   //-------------------------------------------------
   //  Signal enable shot finish
   //-------------------------------------------------
         O(;
   //    u    LastBreakFromExternal    // Signal vom ROBOTER !!!
         A     "DB123_MH_IO_Signals".MH[4].IN.MH_Status.shotactive_MH;
         );
         ON    "DB704_MH_Value".Mixinghead[4].ShotBreak;
         O     "DB123_MH_IO_Signals".MH[4].IN.MH_Manual_Mode;
         S     "EnableFinishShot_MH04";

   //-------------------------------------------------
   // Signal to reset shotrelease
   //-------------------------------------------------
         ON    "DB123_MH_IO_Signals".MH[4].IN.MH_Status.shotactive_MH;
         O     "EnableFinishShot_MH04";
         A     "DB123_MH_IO_Signals".MH[4].IN.MH_Status.shotdone_MH;
         S     "ShotFinishedModul_MH04";
   //-------------------------------------------------
   // Shot release
   //-------------------------------------------------
         A     "DB619_State_MPart".Mixinghead[1].Mixingheadvalve."04";
         AN    "ShotFinishedModul_MH04";
         AN    "DB009_Faults".Fault_State_Grp_1_M1;
         AN    "DB009_Faults".Faults_FKT_Grp_1_M1;
         JCN   SO04;
         L     2#0000_0001;
         L     #ControlBitShot;
         OW;
         T     #ControlBitShot;
   //-------------------------------------------------
   // Shot without Timer
   //-------------------------------------------------
   SO04: CLR;
         JCN   SW04;
         L     2#0000_0010;
         L     #ControlBitShot;
         OW;
         T     #ControlBitShot;
   //-------------------------------------------------
   // Shot with Timer
   //-------------------------------------------------
   SW04: A     "DB619_State_MPart".Mixinghead[1].Mixingheadvalve."04";
         AN    "ShotFinishedModul_MH04";
         AN    "DB009_Faults".Fault_State_Grp_1_M1;
         AN    "DB009_Faults".Faults_FKT_Grp_1_M1;
         JCN   SP04;
         L     2#0000_0100;
         L     #ControlBitShot;
         OW;
         T     #ControlBitShot;
   //-----------------------------------------------------------------
   // Service / Production
   //-----------------------------------------------------------------
   SP04: NOP   0;
         A(;
         ON    #TempShotWithMaterial_M1;
         ON    "DB619_State_MPart".MH_at_Machine[1]."04";
         );
         A(;
         ON    #TempShotWithMaterial_M2;
         ON    "DB619_State_MPart".MH_at_Machine[2]."04";
         );
         ON    "DB614_MH_State".MH_Status[4].Switch_Service_ON_OFF;
         JCN   RF03;
         L     2#0000_1000;
         L     #ControlBitShot;
         OW;
         T     #ControlBitShot;
   //-----------------------------------------------------------------
   // Spare Bit 4..6
   //-----------------------------------------------------------------

   //-----------------------------------------------------------------
   // Reset faults
   //-----------------------------------------------------------------
   RF04: A     "DB009_Faults".HF_Faults_Quit;
         JCN   FE04;
         L     2#1000_0000;
         L     #ControlBitShot;
         OW;
         T     #ControlBitShot;

   FE04: NOP   0;
   //-----------------------------------------------------------------
   // Write Output MH Status
   //-----------------------------------------------------------------
         L     "PN_Mixinghead".Mixinghead[4].Digital.Address;
         L     4;
         +D;
         SLD   3;
         LAR1;
         L     #ControlBitShot;
         T     PQB [ AR1 , P#0.0 ];
   //*****************************************************************
   // Cleaning Piston control of mixing head
   //*****************************************************************
         O(;
         L     "PN_Mixinghead".Mixinghead[4].ReinigungskolbenDigital.Address;
         L     0;
         ==I;
         );
         ON    "PN_Mixinghead".Mixinghead[4].ReinigungskolbenDigital.Active;
         JC    em04;

         L     0;
         T     #ControlBitCP;
   //-------------------------------------------------
   // Request cleaning piston after shot
   //-------------------------------------------------
         A     "DB619_State_MPart".ShotMa[1].ShotData.CP_AfterShot;
   //    U     "DB704_MH_Value".Mixinghead[4].WithCleaningPiston
         JCN   CF04;
         L     2#0000_0001;
         L     #ControlBitCP;
         OW;
         T     #ControlBitCP;
   //-------------------------------------------------
   // Request cleaning piston with button
   //-------------------------------------------------
   CF04: A     "DB614_MH_State".MH_CleaningPiston[4].CP_valve_selected;
         JCN   CM04;
         L     2#0000_0010;
         L     #ControlBitCP;
         OW;
         T     #ControlBitCP;
   //-------------------------------------------------
   // Break forward time
   //-------------------------------------------------
   CM04: NOP   0;
   //-----------------------------------------------------------------
   // Reset faults
   //-----------------------------------------------------------------
         A     "DB009_Faults".HF_Faults_Quit;
         JCN   FC04;
         L     2#0000_1000;
         L     #ControlBitCP;
         OW;
         T     #ControlBitCP;
   //-------------------------------------------------
   FC04: NOP   0;
   //-------------------------------------------------
   // Write Output CP Status
   //-------------------------------------------------
         L     "PN_Mixinghead".Mixinghead[4].ReinigungskolbenDigital.Address;
         SLD   3;
         LAR1;
         L     #ControlBitCP;
         T     PQB [ AR1 , P#0.0 ];
   //-------------------------------------------------
         JU    em04;
   //*****************************************************************
   // Setvalue position of cleaning piston MH 3
   //*****************************************************************
   //      L     "DB896_ConfAnaCP_Contr".AnaCleaningPiston[3].RearPosition
   //      UN    "DB610_State_MPart".Cycle_Ma[1].running
   //      SPB   gap1
   //      L     "DB610_State_MPart".ShotMa[1].ShotValues.CP_ThrottleGap
   //      ITD
   //      DTR
   //      L     "DB604_PV_Mixinghead".Mixinghead[3].CleaningPiston.PV_Conf_ActV.Multiplier
   //      *R
   //      RND
   //      L     "DB604_PV_Mixinghead".Mixinghead[3].CleaningPiston.PV_Conf_ActV.OffsetSignal
   //      ITD
   //      +D
   //gap1: T     #ThrottleGap
   //
   //      L     0
   //      L     "DB1232_ProCanIO_MH".AddressMH[3].Ref_PLC_set_value_CP
   //      <D
   //      SPBN  nz01
   //      SLD   3
   //      LAR1
   //      L     #ThrottleGap
   //      T PAW [ AR1 , P#0.0 ]
   //*****************************************************************
   em04: NOP   0;
END_REGION

REGION Network 11: Mixinghead 5
   //--- mixinghead 5 active at a machine ----------------
         O(;
         L     "DB619_State_MPart".ShotMa[1].ShotData.MH_No;
         L     5;
         ==I;
         );
         O(;
         L     "DB619_State_MPart".ShotMa[2].ShotData.MH_No;
         L     5;
         ==I;
         );
         =     #Temp_MH_Shot_MH05;
         JCN   cr05;

         L     "DB704_MH_Value".Mixinghead[5].Corrvalue;
         T     #Temp_CorrValue;

   // Shottime correction
   cr05: NOP   0;

   //----------------------------------------------------------------
   // Read Shottime for next shot
   //----------------------------------------------------------------
         O     "DB619_State_MPart".Cycle[1].PressurizeTimeRuns;
         O     "DB619_State_MPart".Cycle[1].CtrlChangeTimeRuns;
         A     #Temp_MH_Shot_MH05;
         =     "F_CycleRunningMH05";  // Read corr Shottime

         A     #Temp_MH_Shot_MH05;
         A     "DB619_State_MPart".SWU[1].SWU_OK;
         JCN   om05;

         A     "DB619_State_MPart".Operationmode[1].Operation;
         AN    "DB619_State_MPart".ShotMa[1].ShotData.ShotDisabled;
         =     #Temp_OperationMode;

         AN    "DB619_State_MPart".Cycle[1].running;
         R     "StopShotCorrMH05";
         A     "DB110_Interf_Program_M1".Bits.Stop_Cycle;
         A     "DB619_State_MPart".Cycle[1].running;
         S     "StopShotCorrMH05";

         O     "StopShotCorrMH05";
         O     "DB009_Faults".Fault_State_Grp_1_M1;
         ON    "DB619_State_MPart".Operationmode[1].Controllvoltage;
   //      ON    "DB123_MH_IO_Signals".MH[4].IN.MH_Status.shotdone_MH
         =     #Temp_Error;

         CALL  "FC215_SHOT_ADJUST"
         ( IN_Cycle_running   := "F_CycleRunningMH05",  // "DB610_State_MPart".Cycle_Ma[1].running
           IN_Shot_running    := "M_ShotActive",  // "DB610_State_MPart".Cycle_Ma[1].ShotRuns
           IN_OP_Mode_foaming := #Temp_OperationMode,  // "DB610_State_MPart".Operationmode_Ma[1].Operation
           IN_Error_GRP_1     := #Temp_Error,  // "M1001_FaultLevel_1"
           IN_Tool_no         := "DB619_State_MPart".ToolMa[1].ToolNo,
           IN_PS_no           := "ShotNoNextMa1",  // "DB610_State_MPart".ShotDataMa[1].ShotNo
           IN_Set_Shottime_DB := "DB606_PV_Machine".Machine[1].ShotTime.PV_SetV.Value,
           IN_Actual_Shottime := "DB606_PV_Machine".Machine[1].ShotTime.PV_ActV.Value,
           IN_Corrvalue       := #Temp_CorrValue,
           IN_DB_Shotadjust   := "DB315_ShotadjustS",
           IN_ShotRelease     := "DB619_State_MPart".Cycle[1].Shotrelease,
           IN_MhManual        := 0,  //"DB123_MH_IO_Signals".MH[4].IN.MH_Manual_Mode
           IO_Correct_factor  := "DB614_MH_State".ShotAdjustMH[5].CorrFact,
           IO_PAD_Shottime    := "DB614_MH_State".ShotAdjustMH[5].FoamingTime_ProCan,
           IO_Modul_activ     := "DB614_MH_State".ShotAdjustMH[5].ShotCorrActive,
           IO_Helpflag        := "DB614_MH_State".ShotAdjustMH[5].HFShotCorr,
           IO_Last_Shottime   := "DB614_MH_State".ShotAdjustMH[5].LastShottime,
           IO_Soll_for_Corr   := "DB614_MH_State".ShotAdjustMH[5].SetValueForCorr,
           IO_AdrCorrF        := "DB614_MH_State".ShotAdjustMH[5].AdrCorrFact,
           IO_TestProgram     := "DB614_MH_State".ShotAdjustMH[5].ShotCorrTest,
           IO_CorrTimeTest    := "DB614_MH_State".ShotAdjustMH[5].CorrTimeTest
         );

   // Write mixinghead data to procan mudule
   //----------------------------------------------------------------------
   // Check if the communication partner is ready for
   // data transfer to ProCan
   // ---------------------------------------------------------------------
   om05: NOP   0;
         AN    "PN_Mixinghead".Mixinghead[5].Digital.Active;
         AN    "PN_Mixinghead".Mixinghead[5].Analog.Active;
         JC    em05;
   //-----------------------------------------------------------------
   // Output signals of mixing head modul 4
   //-----------------------------------------------------------------
         A     "DB123_MH_IO_Signals".MH[5].OUT.MH.V_SWU_MH;
         =     "V_SWU_MH05";
         A     "DB123_MH_IO_Signals".MH[5].OUT.MH.H_Shotcounter_MH;
         =     "H_Shotcounter_MH05";
         A     "DB123_MH_IO_Signals".MH[5].OUT.MH.V_CP_Forward_MH;
         =     "V_CP_Forward_MH05";
         A     "DB123_MH_IO_Signals".MH[5].OUT.MH.H_CP_Back_MH;
         =     "H_CP_Back_MH05";
         A     "DB123_MH_IO_Signals".MH[5].OUT.MH.H_Rel_Foaming_MH;
         =     "H_Rel_Foaming_MH05";
         A     "DB123_MH_IO_Signals".MH[5].OUT.MH.H_HighPressure_MH;
         =     "H_HighPressure_MH05";
         A     "DB123_MH_IO_Signals".MH[5].OUT.MH.K_Fault_MC;
         =     "K_Fault_MC05";
         A     "DB123_MH_IO_Signals".MH[5].OUT.MH.K_ShotEnd_MC;
         =     "K_ShotEnd_MC05";
         A     "DB123_MH_IO_Signals".MH[5].OUT.MH.V_MH;
         =     "V_MH_open_MH05";
         A     "DB123_MH_IO_Signals".MH[5].OUT.MH.V_LowPressure_Circ_MH;
         =     "V_LowPressure_Circ_MH05";

   //------------------------------------------------------------
   //
   //     Activate mixinghead at ProCan  modul
   //
   //------------------------------------------------------------

   //--------------- Mixinghead 5 --------------------------------
         O     #Temp_MH_Shot_MH05;
         JCN   SV05;
   //-----------------------------------------------------------------
   // Transmit calculated shot time to ProCan
   //-----------------------------------------------------------------
         L     0;
         L     "PN_Mixinghead".Mixinghead[5].Digital.Address;
         <>D;
         JCN   SV05;
         SLD   3;
         LAR1;
         L     "DB614_MH_State".ShotAdjustMH[5].FoamingTime_ProCan;
         T     PQD[AR1, P#0.0];
   SV05: NOP   0;

   //*****************************************************************
   // Shot control of mixing head
   //*****************************************************************
         L     0;
         T     #ControlBitShot;
   //--------------------------------------------------
   // Shotcycle finished reset signals
   //--------------------------------------------------
         AN    "DB619_State_MPart".Mixinghead[1].Mixingheadvalve."05";
         R     "ShotFinishedModul_MH05";
         R     "EnableFinishShot_MH05";

   //-------------------------------------------------
   //  Signal enable shot finish
   //-------------------------------------------------
         O(;
   //    u    LastBreakFromExternal    // Signal vom ROBOTER !!!
         A     "DB123_MH_IO_Signals".MH[5].IN.MH_Status.shotactive_MH;
         );
         ON    "DB704_MH_Value".Mixinghead[5].ShotBreak;
         O     "DB123_MH_IO_Signals".MH[5].IN.MH_Manual_Mode;
         S     "EnableFinishShot_MH05";

   //-------------------------------------------------
   // Signal to reset shotrelease
   //-------------------------------------------------
         ON    "DB123_MH_IO_Signals".MH[5].IN.MH_Status.shotactive_MH;
         O     "EnableFinishShot_MH05";
         A     "DB123_MH_IO_Signals".MH[5].IN.MH_Status.shotdone_MH;
         S     "ShotFinishedModul_MH05";
   //-------------------------------------------------
   // Shot release
   //-------------------------------------------------
         A     "DB619_State_MPart".Mixinghead[1].Mixingheadvalve."05";
         AN    "ShotFinishedModul_MH05";
         AN    "DB009_Faults".Fault_State_Grp_1_M1;
         AN    "DB009_Faults".Faults_FKT_Grp_1_M1;
         JCN   SO05;
         L     2#0000_0001;
         L     #ControlBitShot;
         OW;
         T     #ControlBitShot;
   //-------------------------------------------------
   // Shot without Timer
   //-------------------------------------------------
   SO05: CLR;
         JCN   SW05;
         L     2#0000_0010;
         L     #ControlBitShot;
         OW;
         T     #ControlBitShot;
   //-------------------------------------------------
   // Shot with Timer
   //-------------------------------------------------
   SW05: A     "DB619_State_MPart".Mixinghead[1].Mixingheadvalve."05";
         AN    "ShotFinishedModul_MH05";
         AN    "DB009_Faults".Fault_State_Grp_1_M1;
         AN    "DB009_Faults".Faults_FKT_Grp_1_M1;
         JCN   SP05;
         L     2#0000_0100;
         L     #ControlBitShot;
         OW;
         T     #ControlBitShot;
   //-----------------------------------------------------------------
   // Service / Production
   //-----------------------------------------------------------------
   SP05: NOP   0;
         A(;
         ON    #TempShotWithMaterial_M1;
         ON    "DB619_State_MPart".MH_at_Machine[1]."05";
         );
         A(;
         ON    #TempShotWithMaterial_M2;
         ON    "DB619_State_MPart".MH_at_Machine[2]."05";
         );
         ON    "DB614_MH_State".MH_Status[5].Switch_Service_ON_OFF;
         JCN   RF05;
         L     2#0000_1000;
         L     #ControlBitShot;
         OW;
         T     #ControlBitShot;
   //-----------------------------------------------------------------
   // Spare Bit 4..6
   //-----------------------------------------------------------------

   //-----------------------------------------------------------------
   // Reset faults
   //-----------------------------------------------------------------
   RF05: A     "DB009_Faults".HF_Faults_Quit;
         JCN   FE05;
         L     2#1000_0000;
         L     #ControlBitShot;
         OW;
         T     #ControlBitShot;

   FE05: NOP   0;
   //-----------------------------------------------------------------
   // Write Output MH Status
   //-----------------------------------------------------------------
         L     "PN_Mixinghead".Mixinghead[5].Digital.Address;
         L     4;
         +D;
         SLD   3;
         LAR1;
         L     #ControlBitShot;
         T     PQB [ AR1 , P#0.0 ];
   //*****************************************************************
   // Cleaning Piston control of mixing head
   //*****************************************************************
         O(;
         L     "PN_Mixinghead".Mixinghead[5].ReinigungskolbenDigital.Address;
         L     0;
         ==I;
         );
         ON    "PN_Mixinghead".Mixinghead[5].ReinigungskolbenDigital.Active;
         JC    em05;

         L     0;
         T     #ControlBitCP;
   //-------------------------------------------------
   // Request cleaning piston after shot
   //-------------------------------------------------
         A     "DB619_State_MPart".ShotMa[1].ShotData.CP_AfterShot;
   //    U     "DB704_MH_Value".Mixinghead[5].WithCleaningPiston
         JCN   CF03;
         L     2#0000_0001;
         L     #ControlBitCP;
         OW;
         T     #ControlBitCP;
   //-------------------------------------------------
   // Request cleaning piston with button
   //-------------------------------------------------
   CF05: A     "DB614_MH_State".MH_CleaningPiston[5].CP_valve_selected;
         JCN   CM05;
         L     2#0000_0010;
         L     #ControlBitCP;
         OW;
         T     #ControlBitCP;
   //-------------------------------------------------
   // Break forward time
   //-------------------------------------------------
   CM05: NOP   0;
   //-----------------------------------------------------------------
   // Reset faults
   //-----------------------------------------------------------------
         A     "DB009_Faults".HF_Faults_Quit;
         JCN   FC05;
         L     2#0000_1000;
         L     #ControlBitCP;
         OW;
         T     #ControlBitCP;
   //-------------------------------------------------
   FC05: NOP   0;
   //-------------------------------------------------
   // Write Output CP Status
   //-------------------------------------------------
         L     "PN_Mixinghead".Mixinghead[5].ReinigungskolbenDigital.Address;
         SLD   3;
         LAR1;
         L     #ControlBitCP;
         T     PQB [ AR1 , P#0.0 ];
   //-------------------------------------------------
         JU    em05;
   //*****************************************************************
   // Setvalue position of cleaning piston MH 3
   //*****************************************************************
   //      L     "DB896_ConfAnaCP_Contr".AnaCleaningPiston[3].RearPosition
   //      UN    "DB610_State_MPart".Cycle_Ma[1].running
   //      SPB   gap1
   //      L     "DB610_State_MPart".ShotMa[1].ShotValues.CP_ThrottleGap
   //      ITD
   //      DTR
   //      L     "DB604_PV_Mixinghead".Mixinghead[3].CleaningPiston.PV_Conf_ActV.Multiplier
   //      *R
   //      RND
   //      L     "DB604_PV_Mixinghead".Mixinghead[3].CleaningPiston.PV_Conf_ActV.OffsetSignal
   //      ITD
   //      +D
   //gap1: T     #ThrottleGap
   //
   //      L     0
   //      L     "DB1232_ProCanIO_MH".AddressMH[3].Ref_PLC_set_value_CP
   //      <D
   //      SPBN  nz01
   //      SLD   3
   //      LAR1
   //      L     #ThrottleGap
   //      T PAW [ AR1 , P#0.0 ]
   //*****************************************************************
   em05: NOP   0;
END_REGION

REGION Network 12: Mixinghead 6
   //--- mixinghead 6 active at a machine ----------------
         O(;
         L     "DB619_State_MPart".ShotMa[1].ShotData.MH_No;
         L     6;
         ==I;
         );
         O(;
         L     "DB619_State_MPart".ShotMa[2].ShotData.MH_No;
         L     6;
         ==I;
         );
         =     #Temp_MH_Shot_MH06;
         JCN   cr06;

         L     "DB704_MH_Value".Mixinghead[6].Corrvalue;
         T     #Temp_CorrValue;

   // Shottime correction
   cr06: NOP   0;

   //----------------------------------------------------------------
   // Read Shottime for next shot
   //----------------------------------------------------------------
         O     "DB619_State_MPart".Cycle[1].PressurizeTimeRuns;
         O     "DB619_State_MPart".Cycle[1].CtrlChangeTimeRuns;
         A     #Temp_MH_Shot_MH06;
         =     "F_CycleRunningMH06";  // Read corr Shottime

         A     #Temp_MH_Shot_MH06;
         A     "DB619_State_MPart".SWU[1].SWU_OK;
         JCN   om06;

         A     "DB619_State_MPart".Operationmode[1].Operation;
         AN    "DB619_State_MPart".ShotMa[1].ShotData.ShotDisabled;
         =     #Temp_OperationMode;

         AN    "DB619_State_MPart".Cycle[1].running;
         R     "StopShotCorrMH06";
         A     "DB110_Interf_Program_M1".Bits.Stop_Cycle;
         A     "DB619_State_MPart".Cycle[1].running;
         S     "StopShotCorrMH06";

         O     "StopShotCorrMH06";
         O     "DB009_Faults".Fault_State_Grp_1_M1;
         ON    "DB619_State_MPart".Operationmode[1].Controllvoltage;
   //      ON    "DB123_MH_IO_Signals".MH[4].IN.MH_Status.shotdone_MH
         =     #Temp_Error;

         CALL  "FC215_SHOT_ADJUST"
         ( IN_Cycle_running   := "F_CycleRunningMH06",  // "DB610_State_MPart".Cycle_Ma[1].running
           IN_Shot_running    := "M_ShotActive",  // "DB610_State_MPart".Cycle_Ma[1].ShotRuns
           IN_OP_Mode_foaming := #Temp_OperationMode,  // "DB610_State_MPart".Operationmode_Ma[1].Operation
           IN_Error_GRP_1     := #Temp_Error,  // "M1001_FaultLevel_1"
           IN_Tool_no         := "DB619_State_MPart".ToolMa[1].ToolNo,
           IN_PS_no           := "ShotNoNextMa1",  // "DB610_State_MPart".ShotDataMa[1].ShotNo
           IN_Set_Shottime_DB := "DB606_PV_Machine".Machine[1].ShotTime.PV_SetV.Value,
           IN_Actual_Shottime := "DB606_PV_Machine".Machine[1].ShotTime.PV_ActV.Value,
           IN_Corrvalue       := #Temp_CorrValue,
           IN_DB_Shotadjust   := "DB315_ShotadjustS",
           IN_ShotRelease     := "DB619_State_MPart".Cycle[1].Shotrelease,
           IN_MhManual        := 0,  //"DB123_MH_IO_Signals".MH[4].IN.MH_Manual_Mode
           IO_Correct_factor  := "DB614_MH_State".ShotAdjustMH[6].CorrFact,
           IO_PAD_Shottime    := "DB614_MH_State".ShotAdjustMH[6].FoamingTime_ProCan,
           IO_Modul_activ     := "DB614_MH_State".ShotAdjustMH[6].ShotCorrActive,
           IO_Helpflag        := "DB614_MH_State".ShotAdjustMH[6].HFShotCorr,
           IO_Last_Shottime   := "DB614_MH_State".ShotAdjustMH[6].LastShottime,
           IO_Soll_for_Corr   := "DB614_MH_State".ShotAdjustMH[6].SetValueForCorr,
           IO_AdrCorrF        := "DB614_MH_State".ShotAdjustMH[6].AdrCorrFact,
           IO_TestProgram     := "DB614_MH_State".ShotAdjustMH[6].ShotCorrTest,
           IO_CorrTimeTest    := "DB614_MH_State".ShotAdjustMH[6].CorrTimeTest
         );

   // Write mixinghead data to procan mudule
   //----------------------------------------------------------------------
   // Check if the communication partner is ready for
   // data transfer to ProCan
   // ---------------------------------------------------------------------
   om06: NOP   0;
         AN    "PN_Mixinghead".Mixinghead[6].Digital.Active;
         AN    "PN_Mixinghead".Mixinghead[6].Analog.Active;
         JC    em06;
   //-----------------------------------------------------------------
   // Output signals of mixing head modul 6
   //-----------------------------------------------------------------
         A     "DB123_MH_IO_Signals".MH[6].OUT.MH.V_SWU_MH;
         =     "V_SWU_MH06";
         A     "DB123_MH_IO_Signals".MH[6].OUT.MH.H_Shotcounter_MH;
         =     "H_Shotcounter_MH06";
         A     "DB123_MH_IO_Signals".MH[6].OUT.MH.V_CP_Forward_MH;
         =     "V_CP_Forward_MH06";
         A     "DB123_MH_IO_Signals".MH[6].OUT.MH.H_CP_Back_MH;
         =     "H_CP_Back_MH06";
         A     "DB123_MH_IO_Signals".MH[6].OUT.MH.H_Rel_Foaming_MH;
         =     "H_Rel_Foaming_MH06";
         A     "DB123_MH_IO_Signals".MH[6].OUT.MH.H_HighPressure_MH;
         =     "H_HighPressure_MH06";
         A     "DB123_MH_IO_Signals".MH[6].OUT.MH.K_Fault_MC;
         =     "K_Fault_MC06";
         A     "DB123_MH_IO_Signals".MH[6].OUT.MH.K_ShotEnd_MC;
         =     "K_ShotEnd_MC06";
         A     "DB123_MH_IO_Signals".MH[6].OUT.MH.V_MH;
         =     "V_MH_open_MH06";
         A     "DB123_MH_IO_Signals".MH[6].OUT.MH.V_LowPressure_Circ_MH;
         =     "V_LowPressure_Circ_MH06";

   //------------------------------------------------------------
   //
   //     Activate mixinghead at ProCan  modul
   //
   //------------------------------------------------------------

   //--------------- Mixinghead 6--------------------------------
         O     #Temp_MH_Shot_MH06;
         JCN   SV06;
   //-----------------------------------------------------------------
   // Transmit calculated shot time to ProCan
   //-----------------------------------------------------------------
         L     0;
         L     "PN_Mixinghead".Mixinghead[6].Digital.Address;
         <>D;
         JCN   SV06;
         SLD   3;
         LAR1;
         L     "DB614_MH_State".ShotAdjustMH[6].FoamingTime_ProCan;
         T     PQD[AR1, P#0.0];
   SV06: NOP   0;

   //*****************************************************************
   // Shot control of mixing head
   //*****************************************************************
         L     0;
         T     #ControlBitShot;
   //--------------------------------------------------
   // Shotcycle finished reset signals
   //--------------------------------------------------
         AN    "DB619_State_MPart".Mixinghead[1].Mixingheadvalve."06";
         R     "ShotFinishedModul_MH06";
         R     "EnableFinishShot_MH06";

   //-------------------------------------------------
   //  Signal enable shot finish
   //-------------------------------------------------
         O(;
   //    u    LastBreakFromExternal    // Signal vom ROBOTER !!!
         A     "DB123_MH_IO_Signals".MH[6].IN.MH_Status.shotactive_MH;
         );
         ON    "DB704_MH_Value".Mixinghead[6].ShotBreak;
         O     "DB123_MH_IO_Signals".MH[6].IN.MH_Manual_Mode;
         S     "EnableFinishShot_MH06";

   //-------------------------------------------------
   // Signal to reset shotrelease
   //-------------------------------------------------
         ON    "DB123_MH_IO_Signals".MH[6].IN.MH_Status.shotactive_MH;
         O     "EnableFinishShot_MH06";
         A     "DB123_MH_IO_Signals".MH[6].IN.MH_Status.shotdone_MH;
         S     "ShotFinishedModul_MH06";
   //-------------------------------------------------
   // Shot release
   //-------------------------------------------------
         A     "DB619_State_MPart".Mixinghead[1].Mixingheadvalve."06";
         AN    "ShotFinishedModul_MH06";
         AN    "DB009_Faults".Fault_State_Grp_1_M1;
         AN    "DB009_Faults".Faults_FKT_Grp_1_M1;
         JCN   SO06;
         L     2#0000_0001;
         L     #ControlBitShot;
         OW;
         T     #ControlBitShot;
   //-------------------------------------------------
   // Shot without Timer
   //-------------------------------------------------
   SO06: CLR;
         JCN   SW06;
         L     2#0000_0010;
         L     #ControlBitShot;
         OW;
         T     #ControlBitShot;
   //-------------------------------------------------
   // Shot with Timer
   //-------------------------------------------------
   SW06: A     "DB619_State_MPart".Mixinghead[1].Mixingheadvalve."06";
         AN    "ShotFinishedModul_MH06";
         AN    "DB009_Faults".Fault_State_Grp_1_M1;
         AN    "DB009_Faults".Faults_FKT_Grp_1_M1;
         JCN   SP06;
         L     2#0000_0100;
         L     #ControlBitShot;
         OW;
         T     #ControlBitShot;
   //-----------------------------------------------------------------
   // Service / Production
   //-----------------------------------------------------------------
   SP06: NOP   0;
         A(;
         ON    #TempShotWithMaterial_M1;
         ON    "DB619_State_MPart".MH_at_Machine[1]."06";
         );
         A(;
         ON    #TempShotWithMaterial_M2;
         ON    "DB619_State_MPart".MH_at_Machine[2]."06";
         );
         ON    "DB614_MH_State".MH_Status[6].Switch_Service_ON_OFF;
         JCN   RF03;
         L     2#0000_1000;
         L     #ControlBitShot;
         OW;
         T     #ControlBitShot;
   //-----------------------------------------------------------------
   // Spare Bit 4..6
   //-----------------------------------------------------------------

   //-----------------------------------------------------------------
   // Reset faults
   //-----------------------------------------------------------------
   RF06: A     "DB009_Faults".HF_Faults_Quit;
         JCN   FE06;
         L     2#1000_0000;
         L     #ControlBitShot;
         OW;
         T     #ControlBitShot;

   FE06: NOP   0;
   //-----------------------------------------------------------------
   // Write Output MH Status
   //-----------------------------------------------------------------
         L     "PN_Mixinghead".Mixinghead[6].Digital.Address;
         L     4;
         +D;
         SLD   3;
         LAR1;
         L     #ControlBitShot;
         T     PQB [ AR1 , P#0.0 ];
   //*****************************************************************
   // Cleaning Piston control of mixing head
   //*****************************************************************
         O(;
         L     "PN_Mixinghead".Mixinghead[3].ReinigungskolbenDigital.Address;
         L     0;
         ==I;
         );
         ON    "PN_Mixinghead".Mixinghead[6].ReinigungskolbenDigital.Active;
         JC    em03;

         L     0;
         T     #ControlBitCP;
   //-------------------------------------------------
   // Request cleaning piston after shot
   //-------------------------------------------------
         A     "DB619_State_MPart".ShotMa[1].ShotData.CP_AfterShot;
   //    U     "DB704_MH_Value".Mixinghead[6].WithCleaningPiston
         JCN   CF06;
         L     2#0000_0001;
         L     #ControlBitCP;
         OW;
         T     #ControlBitCP;
   //-------------------------------------------------
   // Request cleaning piston with button
   //-------------------------------------------------
   CF06: A     "DB614_MH_State".MH_CleaningPiston[6].CP_valve_selected;
         JCN   CM06;
         L     2#0000_0010;
         L     #ControlBitCP;
         OW;
         T     #ControlBitCP;
   //-------------------------------------------------
   // Break forward time
   //-------------------------------------------------
   CM06: NOP   0;
   //-----------------------------------------------------------------
   // Reset faults
   //-----------------------------------------------------------------
         A     "DB009_Faults".HF_Faults_Quit;
         JCN   FC06;
         L     2#0000_1000;
         L     #ControlBitCP;
         OW;
         T     #ControlBitCP;
   //-------------------------------------------------
   FC06: NOP   0;
   //-------------------------------------------------
   // Write Output CP Status
   //-------------------------------------------------
         L     "PN_Mixinghead".Mixinghead[6].ReinigungskolbenDigital.Address;
         SLD   3;
         LAR1;
         L     #ControlBitCP;
         T     PQB [ AR1 , P#0.0 ];
   //-------------------------------------------------
         JU    em06;
   //*****************************************************************
   // Setvalue position of cleaning piston MH 3
   //*****************************************************************
   //      L     "DB896_ConfAnaCP_Contr".AnaCleaningPiston[3].RearPosition
   //      UN    "DB610_State_MPart".Cycle_Ma[1].running
   //      SPB   gap1
   //      L     "DB610_State_MPart".ShotMa[1].ShotValues.CP_ThrottleGap
   //      ITD
   //      DTR
   //      L     "DB604_PV_Mixinghead".Mixinghead[3].CleaningPiston.PV_Conf_ActV.Multiplier
   //      *R
   //      RND
   //      L     "DB604_PV_Mixinghead".Mixinghead[3].CleaningPiston.PV_Conf_ActV.OffsetSignal
   //      ITD
   //      +D
   //gap1: T     #ThrottleGap
   //
   //      L     0
   //      L     "DB1232_ProCanIO_MH".AddressMH[3].Ref_PLC_set_value_CP
   //      <D
   //      SPBN  nz01
   //      SLD   3
   //      LAR1
   //      L     #ThrottleGap
   //      T PAW [ AR1 , P#0.0 ]
   //*****************************************************************
   em06: NOP   0;
END_REGION
END_FUNCTION

FUNCTION "FC205_Tempering_1" : Void   // FC205, STL
TITLE = Heating and cooling depending of the mode
{ S7_Optimized_Access := 'FALSE' }
AUTHOR : KT242
NAME : Temp
VERSION : 2.2
   VAR_INPUT
      IN_Exist : Bool;   // Tempering exist
      IN_Release : Bool;   // Release tempering
      IN_FLT_Ackn : Bool;   // Fault acknowledge
      IN_actual_Temp : Real;
      IN_set_Temp : Real;
   END_VAR
   VAR_IN_OUT
      IO_State : "UDT105_ControllerHeating";   // Controller State of Controller 1
      IO_Values : "UDT702_HeatingControl";   // Values of Controller 1
      IO_Faults : "UDT1804_FLT_Controller";   // Fault bits of Controller 1
      IO_NewFault : Bool;
      IO_FaultLevel_3 : Bool;
   END_VAR
   VAR_TEMP
      Temp_No_Valid_HeatValue : Bool;
      Temp_No_Settings_Requested : Bool;
      Temp_Heating_ON : Real;
      Temp_Heating_OFF : Real;
   END_VAR
BEGIN

REGION Network 1: Relais heating or cooling
         A     #IN_Exist;
         JC    strt;
         R     #IO_State.OUTHeating;
         R     #IO_State.HeatingRequest;
         R     #IO_State.HeatingActive;
         R     #IO_State.Fault_Exist;

         R     #IO_Faults.HW_Limit;
         R     #IO_Faults.Fuse_TemperingOverLoad;
         R     #IO_Faults.lower_limit;
         R     #IO_Faults.upper_limit;
         R     #IO_Faults.NoSetValue;
         BEU;
   strt: NOP   0;
END_REGION

REGION Network 2: Error handling
         A     #IN_FLT_Ackn;
         R     #IO_Faults.HW_Limit;
         R     #IO_Faults.Fuse_TemperingOverLoad;
         R     #IO_Faults.lower_limit;
         R     #IO_Faults.upper_limit;
         R     #IO_Faults.NoSetValue;

   // Sets fault if man.temp > 0 and act.temp > max.temp
         A(;
         L     #IO_Values.Max_Temp;
         L     0.0;
         >R;
         );
         A(;
         L     #IN_actual_Temp;
         L     #IO_Values.Max_Temp;
         >R;
         );
         A     #IO_State.Switch_ON_OFF;
         AN    #IO_Faults.upper_limit;
         S     #IO_NewFault;
         S     #IO_Faults.upper_limit;

         AN    #IO_State.INFuse;
         A     #IO_State.Switch_ON_OFF;
         AN    #IO_Faults.Fuse_TemperingOverLoad;
         S     #IO_NewFault;
         S     #IO_Faults.Fuse_TemperingOverLoad;

         A     #IO_State.INHeatingLimit;
         A     #IO_State.Switch_ON_OFF;
         AN    #IO_Faults.HW_Limit;
         S     #IO_NewFault;
         S     #IO_Faults.HW_Limit;

         A(;
         L     #IN_set_Temp;
         L     0.0;
         ==R;
         );
         A     #IO_State.Switch_ON_OFF;
         AN    #IO_Faults.NoSetValue;
         S     #IO_NewFault;
         S     #IO_Faults.NoSetValue;

         O     #IO_Faults.HW_Limit;
         O     #IO_Faults.Fuse_TemperingOverLoad;
         O     #IO_Faults.lower_limit;
         O     #IO_Faults.upper_limit;
         O     #IO_Faults.NoSetValue;
         O     #IO_Faults.Sensor_FLT_broken_wire;
         O     #IO_Faults.Warning_limit_plus;
         O     #IO_Faults.Warning_limit_minus;
         O     #IO_Faults.Alarm_limit_plus;
         O     #IO_Faults.Alarm_limit_minus;
         O     #IO_Faults.Controller_at_limit;
         S     #IO_FaultLevel_3;
         =     #IO_State.Fault_Exist;
END_REGION

REGION Network 3: Test the values
         O(;
         L     #IO_Values.Dif_Heating_ON;
         L     0.0;
         ==R;
         );
         O(;
         L     #IO_Values.Dif_Heating_ON;
         L     #IO_Values.Dif_Heating_OFF;
         <R;
         );
         =     #Temp_No_Valid_HeatValue;
END_REGION

REGION Network 4: Calculate limits
         L     #IN_set_Temp;
         L     #IO_Values.Dif_Heating_ON;
         -R;
         T     #Temp_Heating_ON;

         L     #IN_set_Temp;
         L     #IO_Values.Dif_Heating_OFF;
         -R;
         T     #Temp_Heating_OFF;
END_REGION

REGION Network 5: Heating mode
   // Kühlen ist dominant
         O     #IO_Faults.NoSetValue;
         R     #IO_State.HeatingRequest;
         JC    OUTH;

         L     #IN_actual_Temp;  // Actual Temp < Switch ON value
         L     #Temp_Heating_ON;
         <R;
         S     #IO_State.HeatingRequest;

         A(;
         L     #IN_actual_Temp;
         L     #IO_Values.Max_Temp;
         >R;
         );
         A(;
         L     #IO_Values.Max_Temp;
         L     0.0;
         >R;
         );
         O(;
         L     #IN_actual_Temp;
         L     #Temp_Heating_OFF;
         >=R;
         );
         O     #Temp_No_Valid_HeatValue;
         ON    #IO_State.Switch_ON_OFF;
         R     #IO_State.HeatingRequest;

   OUTH: NOP   0;

         A     #IN_Exist;
         A     #IN_Release;
         A     #IO_State.HeatingRequest;
         AN    #IO_Faults.Fuse_TemperingOverLoad;
         AN    #IO_Faults.HW_Limit;
         AN    #IO_Faults.upper_limit;
         =     #IO_State.OUTHeating;
         =     #IO_State.HeatingActive;
END_REGION

REGION Network 6: State tempering 1: ON; 2:error; 3:Selected but not ON
         L     0;
         O     #IO_Faults.Fuse_TemperingOverLoad;
         O     #IO_Faults.HW_Limit;
         JCN   F_ON;
         L     2;
         JU    tran;
   F_ON: O     #IO_State.HeatingActive;
         JCN   anl;
         L     1;
         JU    tran;
   anl:  ON    #IO_State.Switch_ON_OFF;
         O     #IO_State.HeatingActive;
         JC    tran;
         L     3;
   tran: T     #IO_State.State_Temp;
END_REGION
END_FUNCTION

FUNCTION "FC215_SHOT_ADJUST" : Void   // FC215, STL
TITLE = Shottime adjustment
{ S7_Optimized_Access := 'FALSE' }
AUTHOR : HK
NAME : ShotTime
VERSION : 0.4
   VAR_INPUT
      IN_Cycle_running : Bool;
      IN_Shot_running : Bool;
      IN_OP_Mode_foaming : Bool;
      IN_Error_GRP_1 : Bool;
      IN_Tool_no : Int;   // Number of tool
      IN_PS_no : Int;   // Part shot number
      IN_Set_Shottime_DB : Real;   // Set shot time
      IN_Actual_Shottime : Real;   // actual shot time
      IN_Corrvalue : Real;   // Factor runtime steering piston
      IN_DB_Shotadjust : DB_ANY;
      IN_ShotRelease : Bool;
      IN_MhManual : Bool;   // Mixinghead in manual -> Testshot selected
   END_VAR
   VAR_IN_OUT
      IO_Correct_factor : Real;   // Corrrction factor
      IO_PAD_Shottime : Real;   // Address of corr shot time
      IO_Modul_activ : Bool;   // Modul is active
      IO_Helpflag : Bool;
      IO_Last_Shottime : Real;
      IO_Soll_for_Corr : Real;
      IO_AdrCorrF : DWord;
      IO_TestProgram : Bool;   // Test program is running - dont't write correction time to DB
      IO_CorrTimeTest : Real;   // Correcting time for test shots
   END_VAR
   VAR_TEMP
      Temp_Startaddress : Word;
      Temp_Offset : Word;
      Temp_Poi_ok : Bool;
      Temp_Adr_Corr : DWord;
      TempCorrFactor : Real;
   END_VAR
BEGIN

REGION Network 1: Shottime adjustment max. value 250 ms; limit toolno. partshot no
         O(;
         L     #IO_Correct_factor;
         L     0.25;
         >R;
         );
         O(;
         L     #IO_Correct_factor;
         L     -0.25;
         <R;
         );
         JCN   NW1E;
   ///
         L     0.061;
         T     #IO_Correct_factor;
   ///
   NW1E: NOP   0;

   // Zeiger gültig?
         L     #IN_Tool_no;
         L     0;
         <>I;
         A(;
         L     #IN_Tool_no;
         L     255;
         <=I;
         );
         A(;
         L     #IN_PS_no;
         L     0;
         <>I;
         );
         A(;
         L     #IN_PS_no;
         L     32;
         <=I;
         );
         =     #Temp_Poi_ok;


         AN    #Temp_Poi_ok;
         BEC;
END_REGION

REGION Network 2: Calculate shottime to transfer at Procan modul
         ON    #IN_Cycle_running;
         O(;
         L     #IN_Tool_no;
         L     0;
         ==I;
         );
         O(;
         L     #IN_PS_no;
         L     0;
         ==I;
         );
         R     #IO_TestProgram;
         JC    NW2E;
   ///
         A     #IN_Cycle_running;
         A     #IN_MhManual;
         S     #IO_TestProgram;
   ///
   // Calculate pointer at correction value
         A     #IO_TestProgram;
         JC    ldt;  // load test data

         L     #IN_Tool_no;  // No. of actual used tool
         L     8;  // Amount of partshots per tool
         *D;
         T     #Temp_Startaddress;  // Startaddress at DB of 1. partshot

         L     #IN_PS_no;
         L     1;
         -D;
         T     #Temp_Offset;

         L     #Temp_Startaddress;  // Anfangsadresse im Programm-DB für 1. Teilschuss
         L     #Temp_Offset;  // Offset für 2./3./4. Teilschuss berechnen
         +D;
         SLD   4;  // Adresse im DB
         A     #IN_ShotRelease;
         SET;
         JCN   corr;
         T     #IO_AdrCorrF;
   corr: L     #IO_AdrCorrF;
         LAR2;
         OPN   #IN_DB_Shotadjust;
         L     DBD [ AR2 , P#0.0 ];
         JU    crr;
   ldt:  L     #IO_CorrTimeTest;
   crr:  T     #IO_Correct_factor;  // Ist jetzt Speicher für letzte Korrektur

   // Nochmal limitieren, weil ja erst hier geholt wird !!!
         O(;
         L     #IO_Correct_factor;
         L     0.25;
         >R;
         );
         O(;
         L     #IO_Correct_factor;
         L     -0.25;
         <R;
         );
         JCN   tr;
   ///
         L     0.061;
         T     #IO_Correct_factor;
   ///
   tr:   A     #IN_OP_Mode_foaming;  // bei Service keine Schusszeitkorrektur
         L     #IN_Set_Shottime_DB;
         JCN   SHT;
   ///
         L     #IO_Correct_factor;  // Schusszeitkorrektur
         T     #TempCorrFactor;

         L     #IN_Set_Shottime_DB;
         L     #TempCorrFactor;  // Schusszeitkorrektur
         -R;
         L     #IN_Corrvalue;  // ab V0.2
         -R;
   ///
   SHT:  NOP   0;
         T     #IO_PAD_Shottime;  // Schusszeit an Ausgangsdoppelwort
   NW2E: NOP   0;
END_REGION

REGION Network 3: Calculate correction factor
         A     #IN_Shot_running;
         S     #IO_Modul_activ;  // Modul is active
   ///
         A     #IN_Shot_running;  // Sollwert für Korrektur erst bei Schussbeginn übernehmen
         JCN   keKo;
         L     #IN_Set_Shottime_DB;
         T     #IO_Soll_for_Corr;
   keKo: NOP   0;

         A     #IN_Shot_running;
         A     #IO_Modul_activ;
         FN    #IO_Helpflag;
         JCN   NW3E;
   ///
         L     #IN_Actual_Shottime;
         T     #IO_Last_Shottime;
         AN    #IN_OP_Mode_foaming;
         JC    nc;
         L     #IN_Corrvalue;
         +R;
         T     #IO_Last_Shottime;
   ///
   nc:   SET;
         R     #IO_Modul_activ;  // Modul ist aktiv
   ///
         O     #IN_Error_GRP_1;
         ON    #IN_OP_Mode_foaming;
         JC    NW3E;
   ///
         L     #IO_Last_Shottime;
         L     #IO_Soll_for_Corr;
         -R;
         L     #IO_Correct_factor;
         +R;
         T     #IO_Correct_factor;

         A     #IO_TestProgram;
         JC    crts;

         L     #IO_AdrCorrF;
         LAR2;
         OPN   #IN_DB_Shotadjust;
         L     #IO_Correct_factor;  // Ist jetzt Speicher für letzte Korrektur
         T     DBD [ AR2 , P#0.0 ];
         JU    NW3E;

   crts: L     #IO_Correct_factor;
         T     #IO_CorrTimeTest;
   ///
   NW3E: NOP   0;
END_REGION
END_FUNCTION

FUNCTION "FC216_2-point_adjust" : Void   // FC216, SCL
{ S7_Optimized_Access := 'TRUE' }
VERSION : 0.1
   VAR_TEMP
      Ti_Loop_pump : Int;
   END_VAR
BEGIN
   // Selection for 2 point adjust
   // Use set values for the pump (Don't use QPB values)

   FOR #Ti_Loop_pump := 1 TO 8 DO
       IF "DB613_Komponent_State".MeteringPump[#Ti_Loop_pump].Metering_to_PUC THEN
           IF ("DB613_Komponent_State".FlowPump[#Ti_Loop_pump] > "DB753_MeteringPump".Pump[#Ti_Loop_pump].FlowThreshold) AND "DB753_MeteringPump".Pump[#Ti_Loop_pump].With_2Point THEN
               "DB613_Komponent_State".MeteringPump[#Ti_Loop_pump]."2PointAdjustmentSelected" := True;
           ELSE
               "DB613_Komponent_State".MeteringPump[#Ti_Loop_pump]."2PointAdjustmentSelected" := false;
           END_IF;
       END_IF;
   END_FOR;

   // If version with selection in the mould editor is used, uncomment the rows for "2PointAdjustmentSelected" in FC1156 (6x) and activate in FB4 ( "InterfaceVisu"."2PoinMovementComp"[#TiLoop_Flow]) and don't use this FC
END_FUNCTION

FUNCTION "FC217_Calc_flow_limits" : Void   // FC217, SCL
{ S7_Optimized_Access := 'TRUE' }
VERSION : 0.1
// Calculate min and max value flow for pumps
   VAR_TEMP
      Ti_tank : Int;
      Ti_comp : Int;
      tank_no : Int;   // tank number of pump
      MaxFlowPump : Real;   // Max flow in cm³/s
   END_VAR
BEGIN
   // Density: g/l
   // MaxFlowPump: cm³/s
   // MaxFlowLiter: l
   // FlowPumpMin: g/s
   // FlowPumpMax: g/s

   REGION Calculate the minimum/maximum flow rate of the pumps
       FOR #Ti_comp := 0 TO 12 DO
           #tank_no := "DB753_MeteringPump".Pump[#Ti_comp].TankNo;
           IF #tank_no <> 0 THEN
               #MaxFlowPump := "DB753_MeteringPump".Pump[#Ti_comp].MaxFlowLiter / 0.06;
               "DB613_Komponent_State".FlowPumpMin[#Ti_comp] := ((INT_TO_REAL("DB702_Tank_Value".Tank[#tank_no].Density) / 1000.0) * #MaxFlowPump) / 100 * "DB753_MeteringPump".Pump[#Ti_comp].MinFlowPercent;
               "DB613_Komponent_State".FlowPumpMax[#Ti_comp] := ((INT_TO_REAL("DB702_Tank_Value".Tank[#tank_no].Density) / 1000.0) * #MaxFlowPump) / 100 * "DB753_MeteringPump".Pump[#Ti_comp].MaxFlowPercent;
           END_IF;
       END_FOR;
   END_REGION
END_FUNCTION

FUNCTION "FC916_PV_Limits" : Void   // FC916, STL
TITLE = Checks the limits of a process value
{ S7_Optimized_Access := 'FALSE' }
VERSION : 0.1
   VAR_INPUT
      IN_Tolerance_Test : Bool;
      IN_Reset_Fault : Bool;
   END_VAR
   VAR_IN_OUT
      IO_Any_ArrayPV : ANY;
      IO_Fault_Warn_upperL : Bool;
      IO_Fault_Warn_lowerL : Bool;
      IO_Fault_Alarm_upperL : Bool;
      IO_Fault_Alarm_lowerL : Bool;
      IO_New_Fault : Bool;
      IO_Fault_Level_1 : Bool;
      IO_Fault_Level_2 : Bool;
      IO_Fault_Level_3 : Bool;
   END_VAR
   VAR_TEMP
      RetVal : Int;
      Anf_DW_PV_Act : Word;
      Anyzeiger_PV : ANY;
      Temp_PV : "UDT910_ProcessValue";
      Temp_Counter_average_r : DWord;
      Temp_ActV_Pointer : DWord;
   END_VAR
BEGIN

REGION Network 2: Read Array[No_Array] actual value and set value
         L;  // Pointer auf erstes Element des Arrays
         LAR1;

         LAR2;
   //
         L     W[AR1, P#0.0];  // Bytes
         T     W[AR2, P#0.0];
         L     W [ AR1 , P#2.0 ];  // Amount of bytes
         T     W[AR2, P#2.0];
         L     W [ AR1 , P#4.0 ];  // Block no,
         T     W[AR2, P#4.0];
         L     D [ AR1 , P#6.0 ];  // Startadress of datas
         T     D[AR2, P#6.0];
   //

         CALL  BLKMOV
         ( SRCBLK  := #Anyzeiger_PV,
           RET_VAL := #RetVal,
           DSTBLK  := #Temp_PV
         );
   //
END_REGION

REGION Network 3
   //-----------------------------------------------
   // Alarm limit below
   //-----------------------------------------------
         AN    #IN_Reset_Fault;
         JC    n011;
         L     0;
         T     #Temp_PV.PV_ActV.ValueState;

         R     #IO_Fault_Alarm_lowerL;
         R     #IO_Fault_Alarm_upperL;

         R     #IO_Fault_Warn_lowerL;
         R     #IO_Fault_Warn_upperL;

   n011: A     #IN_Tolerance_Test;
         JC    n012;
         L     0;
         T     #Temp_PV.PV_ActV.ValueState;

         JC    ENDC;

   n012: O(;
         L     #Temp_PV.PV_SetV.AlarmLowerLimit;
         L     0.0;
         <=R;
         );
         O(;
         L     #Temp_PV.PV_SetV.Value;
         L     #Temp_PV.PV_SetV.AlarmLowerLimit;
         -R;
         L     #Temp_PV.PV_ActV.Value;
         <R;
         );
         JC    alun;

         L     1;
         T     #Temp_PV.PV_ActV.ValueState;

         JU    end;

   alun: NOP   0;

   //-----------------------------------------------
   // Warning limit lower
   //-----------------------------------------------
         O(;
         L     #Temp_PV.PV_SetV.WarningLowerLimit;
         L     0.0;
         <=R;
         );
         O(;
         L     #Temp_PV.PV_SetV.Value;
         L     #Temp_PV.PV_SetV.WarningLowerLimit;
         -R;
         L     #Temp_PV.PV_ActV.Value;
         <R;
         );
         JC    gwun;

         L     2;
         T     #Temp_PV.PV_ActV.ValueState;

         JU    end;

   gwun: NOP   0;

         O(;
         L     #Temp_PV.PV_SetV.AlarmUpperLimit;
         L     0.0;
         <=R;
         );
         O(;
         L     #Temp_PV.PV_SetV.Value;
         L     #Temp_PV.PV_SetV.AlarmUpperLimit;
         +R;
         L     #Temp_PV.PV_ActV.Value;
         >R;
         );
         JC    alon;

         L     8;
         T     #Temp_PV.PV_ActV.ValueState;

         JU    end;

   alon: NOP   0;